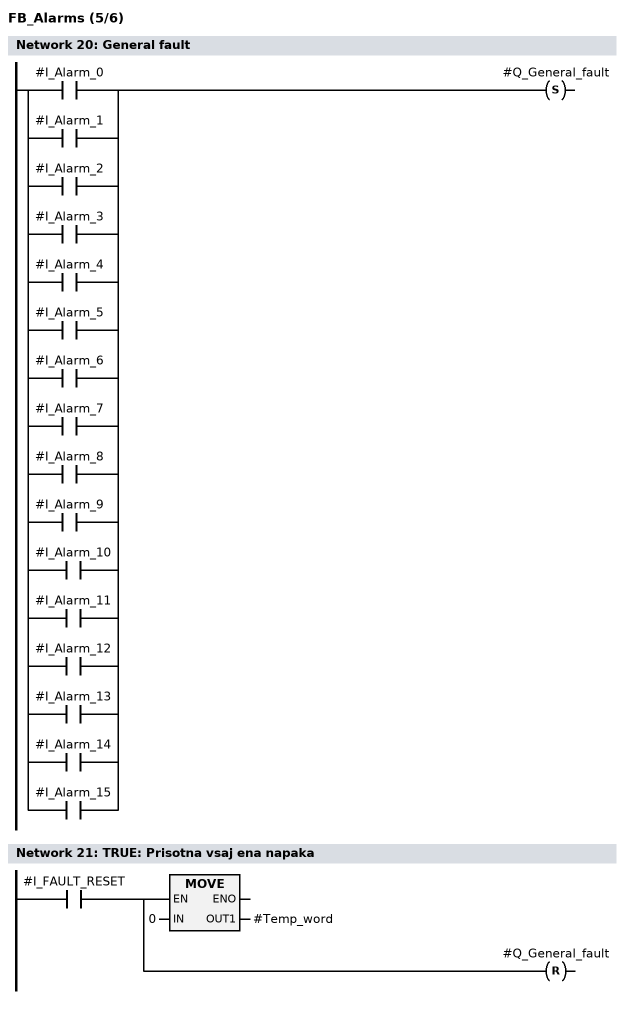
   RUNG wire#powerrail
      Contact( #I_Alarm_0 )
      wire#w1
      S_Coil( #Q_General_fault )
   END_RUNG
   RUNG wire#powerrail
      Contact( #I_Alarm_1 )
   END_RUNG wire#w1
   RUNG wire#powerrail
      Contact( #I_Alarm_2 )
   END_RUNG wire#w1
   RUNG wire#powerrail
      Contact( #I_Alarm_3 )
   END_RUNG wire#w1
   RUNG wire#powerrail
      Contact( #I_Alarm_4 )
   END_RUNG wire#w1
   RUNG wire#powerrail
      Contact( #I_Alarm_5 )
   END_RUNG wire#w1
   RUNG wire#powerrail
      Contact( #I_Alarm_6 )
   END_RUNG wire#w1
   RUNG wire#powerrail
      Contact( #I_Alarm_7 )
   END_RUNG wire#w1
   RUNG wire#powerrail
      Contact( #I_Alarm_8 )
   END_RUNG wire#w1
   RUNG wire#powerrail
      Contact( #I_Alarm_9 )
   END_RUNG wire#w1
   RUNG wire#powerrail
      Contact( #I_Alarm_10 )
   END_RUNG wire#w1
   RUNG wire#powerrail
      Contact( #I_Alarm_11 )
   END_RUNG wire#w1
   RUNG wire#powerrail
      Contact( #I_Alarm_12 )
   END_RUNG wire#w1
   RUNG wire#powerrail
      Contact( #I_Alarm_13 )
   END_RUNG wire#w1
   RUNG wire#powerrail
      Contact( #I_Alarm_14 )
   END_RUNG wire#w1
   RUNG wire#powerrail
      Contact( #I_Alarm_15 )
   END_RUNG wire#w1
   // the same network as SCL:
   IF #I_Alarm_0 OR #I_Alarm_1 OR #I_Alarm_2 OR #I_Alarm_3 OR #I_Alarm_4 OR #I_Alarm_5 OR #I_Alarm_6 OR #I_Alarm_7 OR #I_Alarm_8 OR #I_Alarm_9 OR #I_Alarm_10 OR #I_Alarm_11 OR #I_Alarm_12 OR #I_Alarm_13 OR #I_Alarm_14 OR #I_Alarm_15 THEN
       #Q_General_fault := TRUE;
   END_IF;
END_REGION

REGION Network 21: TRUE: Prisotna vsaj ena napaka
   RUNG wire#powerrail
      Contact( #I_FAULT_RESET )
      wire#w1
      { S7_GenerateENO := "TRUE" } Move(in := 0, out1 => #Temp_word)
   END_RUNG
   RUNG wire#w1
      R_Coil( #Q_General_fault )
   END_RUNG
   // the same network as SCL:
   IF #I_FAULT_RESET THEN
       #Temp_word := 0;
       #Q_General_fault := FALSE;
   END_IF;
END_REGION

REGION Network 23
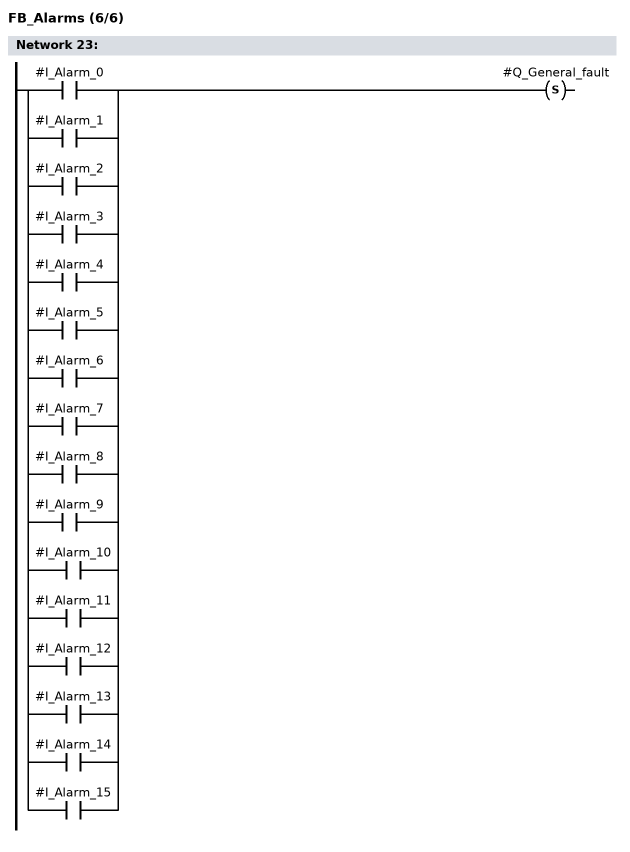
   RUNG wire#powerrail
      Contact( #I_Alarm_0 )
      wire#w1
      S_Coil( #Q_General_fault )
   END_RUNG
   RUNG wire#powerrail
      Contact( #I_Alarm_1 )
   END_RUNG wire#w1
   RUNG wire#powerrail
      Contact( #I_Alarm_2 )
   END_RUNG wire#w1
   RUNG wire#powerrail
      Contact( #I_Alarm_3 )
   END_RUNG wire#w1
   RUNG wire#powerrail
      Contact( #I_Alarm_4 )
   END_RUNG wire#w1
   RUNG wire#powerrail
      Contact( #I_Alarm_5 )
   END_RUNG wire#w1
   RUNG wire#powerrail
      Contact( #I_Alarm_6 )
   END_RUNG wire#w1
   RUNG wire#powerrail
      Contact( #I_Alarm_7 )
   END_RUNG wire#w1
   RUNG wire#powerrail
      Contact( #I_Alarm_8 )
   END_RUNG wire#w1
   RUNG wire#powerrail
      Contact( #I_Alarm_9 )
   END_RUNG wire#w1
   RUNG wire#powerrail
      Contact( #I_Alarm_10 )
   END_RUNG wire#w1
   RUNG wire#powerrail
      Contact( #I_Alarm_11 )
   END_RUNG wire#w1
   RUNG wire#powerrail
      Contact( #I_Alarm_12 )
   END_RUNG wire#w1
   RUNG wire#powerrail
      Contact( #I_Alarm_13 )
   END_RUNG wire#w1
   RUNG wire#powerrail
      Contact( #I_Alarm_14 )
   END_RUNG wire#w1
   RUNG wire#powerrail
      Contact( #I_Alarm_15 )
   END_RUNG wire#w1
   // the same network as SCL:
   IF #I_Alarm_0 OR #I_Alarm_1 OR #I_Alarm_2 OR #I_Alarm_3 OR #I_Alarm_4 OR #I_Alarm_5 OR #I_Alarm_6 OR #I_Alarm_7 OR #I_Alarm_8 OR #I_Alarm_9 OR #I_Alarm_10 OR #I_Alarm_11 OR #I_Alarm_12 OR #I_Alarm_13 OR #I_Alarm_14 OR #I_Alarm_15 THEN
       #Q_General_fault := TRUE;
   END_IF;
END_REGION
END_FUNCTION_BLOCK

FUNCTION_BLOCK "BOOL_TO_INT"   // FB125, LAD
TITLE = Alarm blok
{ S7_Optimized_Access := 'TRUE' }
AUTHOR : Andrej
VERSION : 0.1
   VAR_INPUT
      BOOL_0 : Bool;
      BOOL_1 : Bool;
      BOOL_2 : Bool;
      BOOL_3 : Bool;
      BOOL_4 : Bool;
      BOOL_5 : Bool;
      BOOL_6 : Bool;
      BOOL_7 : Bool;
      BOOL_8 : Bool;
      BOOL_9 : Bool;
      BOOL_10 : Bool;
      BOOL_11 : Bool;
      BOOL_12 : Bool;
      BOOL_13 : Bool;
      BOOL_14 : Bool;
      BOOL_15 : Bool;
   END_VAR
   VAR_OUTPUT
      "INT" : Word;
   END_VAR
   VAR RETAIN
      Temp_word : Word;
   END_VAR
BEGIN

REGION Network 1
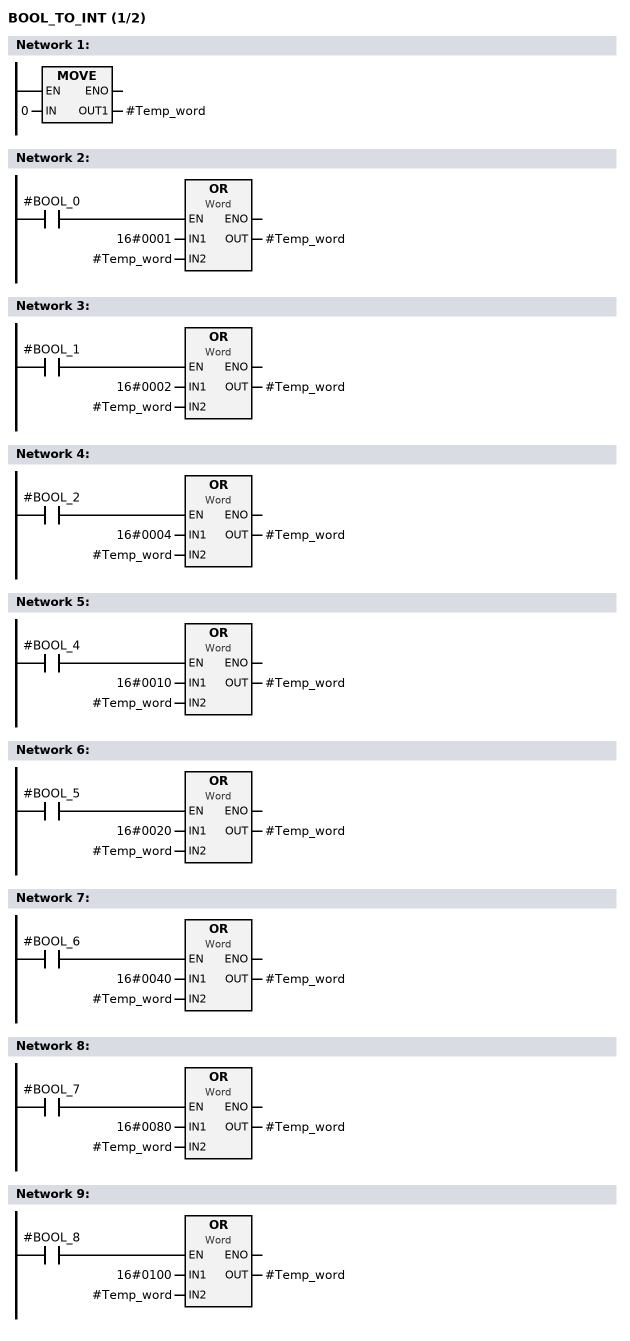
   RUNG wire#powerrail
      Move(in := 0, out1 => #Temp_word)
   END_RUNG
   // the same network as SCL:
   #Temp_word := 0;
END_REGION

REGION Network 2
   IF #BOOL_0 THEN #Temp_word := 16#0001 OR #Temp_word; END_IF;
END_REGION

REGION Network 3
   IF #BOOL_1 THEN #Temp_word := 16#0002 OR #Temp_word; END_IF;
END_REGION

REGION Network 4
   IF #BOOL_2 THEN #Temp_word := 16#0004 OR #Temp_word; END_IF;
END_REGION

REGION Network 5
   IF #BOOL_4 THEN #Temp_word := 16#0010 OR #Temp_word; END_IF;
END_REGION

REGION Network 6
   IF #BOOL_5 THEN #Temp_word := 16#0020 OR #Temp_word; END_IF;
END_REGION

REGION Network 7
   IF #BOOL_6 THEN #Temp_word := 16#0040 OR #Temp_word; END_IF;
END_REGION

REGION Network 8
   IF #BOOL_7 THEN #Temp_word := 16#0080 OR #Temp_word; END_IF;
END_REGION

REGION Network 9
   IF #BOOL_8 THEN #Temp_word := 16#0100 OR #Temp_word; END_IF;
END_REGION

REGION Network 10
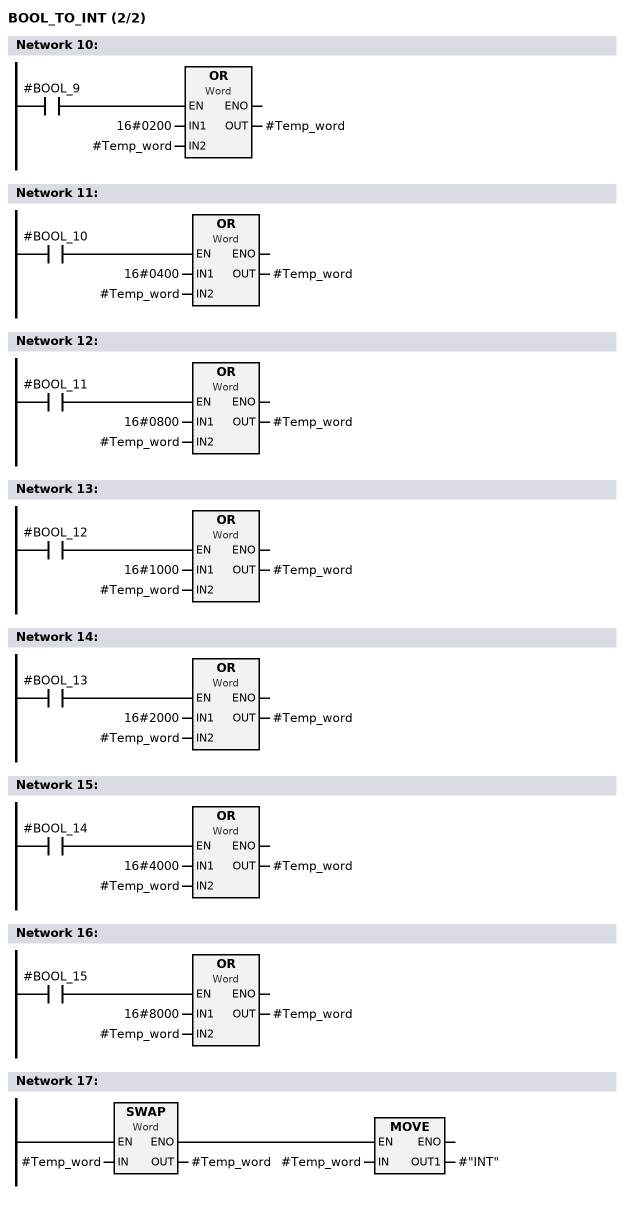
   IF #BOOL_9 THEN #Temp_word := 16#0200 OR #Temp_word; END_IF;
END_REGION

REGION Network 11
   IF #BOOL_10 THEN #Temp_word := 16#0400 OR #Temp_word; END_IF;
END_REGION

REGION Network 12
   IF #BOOL_11 THEN #Temp_word := 16#0800 OR #Temp_word; END_IF;
END_REGION

REGION Network 13
   IF #BOOL_12 THEN #Temp_word := 16#1000 OR #Temp_word; END_IF;
END_REGION

REGION Network 14
   IF #BOOL_13 THEN #Temp_word := 16#2000 OR #Temp_word; END_IF;
END_REGION

REGION Network 15
   IF #BOOL_14 THEN #Temp_word := 16#4000 OR #Temp_word; END_IF;
END_REGION

REGION Network 16
   IF #BOOL_15 THEN #Temp_word := 16#8000 OR #Temp_word; END_IF;
END_REGION

REGION Network 17
   #Temp_word := SWAP(#Temp_word);
   #"INT" := #Temp_word;
END_REGION
END_FUNCTION_BLOCK

(* ===== HMI "HMI_RT_6" =====
system functions are stored by id; their names below are inferred from use
connection "HMI_Connection_8": 
connection "HMI_Connection_1": ETHERNET, S7_1500_OMS

HMI tags "Default tag table"
   "PozKontaktNaKoncuLetve" : Bool = PLC PozKontaktNaKoncuLetve AT %I20.4, 1 s
   "FB_STARTUP_DB_korak" : UInt = PLC FB_STARTUP_DB.korak, 1 s
   "FB_IOL_IFM_SV_DB_uPretok" : UInt = PLC FB_IOL_IFM_SV_DB.uPretok, 1 s
   "FB_IOL_IFM_SV_DB_fTemperatura" : Real = PLC FB_IOL_IFM_SV_DB.fTemperatura, 1 s
   "FB_FESTO_VPPM_DB_TrenutniPritisk" : Real = PLC FB_FESTO_VPPM_DB.TrenutniPritisk, 1 s
   "FB_FESTO_SDE1_DB_oPritisk" : Real = PLC FB_FESTO_SDE1_DB.oPritisk, 1 s
   "FB_Lin_FESTO_PNEVMATIKA_PRITISK_Q_izhod" : Real = PLC FB_Lin_FESTO_PNEVMATIKA_PRITISK.Q_izhod, 1 s
   "FB_FESTO_VPPM_DB_setstatZeljeniPritisk" : Real = PLC FB_FESTO_VPPM_DB.setstatZeljeniPritisk, 1 s
   "Keyence_OdmičniCilinderKonusa" : DInt = PLC Keyence_OdmičniCilinderKonusa AT %ID137, 1 s
   "Keyence_OdmičniCilinderVarjenja" : DInt = PLC Keyence_OdmičniCilinderVarjenja AT %ID144, 1 s
   "DB_HMI_ROČNI NAČIN_izbraniCilinder" : Int = PLC DB_HMI."ROČNI NAČIN".izbraniCilinder, 1 s
   "ZaporaIzdelka" : Bool = PLC ZaporaIzdelka AT %I20.0, 1 s
   "SprositevZaporeIzdelka" : Bool = PLC SprositevZaporeIzdelka AT %I20.1, 1 s
   "1Y1_OdklepZapore" : Bool = PLC 1Y1_OdklepZapore AT %Q44.0, 1 s
   "Y2/1_NalaganjeNazanj" : Bool = PLC "Y2/1_NalaganjeNazanj" AT %Q44.3, 1 s
   "Y2/1_NalaganjeNaprej" : Bool = PLC "Y2/1_NalaganjeNaprej" AT %Q44.2, 1 s
   "DB_HMI_SDAT1_PozPobiranje" : Real = PLC DB_HMI.SDAT1.PozPobiranje, 1 s
   "DB_HMI_SDAT1_PozNalaganje" : Real = PLC DB_HMI.SDAT1.PozNalaganje, 1 s
   "SDAT1_oPoz1Dosezena" : Bool = PLC SDAT1.oPoz1Dosezena, 1 s
   "SDAT2_oPoz2Dosezena" : Bool = PLC SDAT2.oPoz2Dosezena, 1 s
   "SDAT1_oPoz2Dosezena" : Bool = PLC SDAT1.oPoz2Dosezena, 1 s
   "Y3/1_PrijemaloKontaktaOdpri" : Bool = PLC "Y3/1_PrijemaloKontaktaOdpri" AT %Q44.4, 1 s
   "PrijemaloKontaktaOdprto" : Bool = PLC PrijemaloKontaktaOdprto AT %I20.3, 1 s
   "PrijemaloKontaktaZaprto" : Bool = PLC PrijemaloKontaktaZaprto AT %I20.2, 1 s
   "DB_HMI_SDAT2_PozNalaganje" : Real = PLC DB_HMI.SDAT2.PozPobiranjePloscice, 1 s
   "DB_HMI_SDAT2_PozPobiranje" : Real = PLC DB_HMI.SDAT2.PozNalaganjePloscice, 1 s
   "SDAT1_out" : Real = PLC SDAT1.out, 1 s
   "SDAT2_out" : Real = PLC SDAT2.out, 1 s
   "FB_KEYENCE_GT2_ODMIKVARJENJA_oPoz1Dosezena" : Bool = PLC FB_KEYENCE_GT2_ODMIKVARJENJA.oPoz1Dosezena, 1 s
   "FB_KEYENCE_GT2_ODMIKVARJENJA_oPoz3Dosezena" : Bool = PLC FB_KEYENCE_GT2_ODMIKVARJENJA.oPoz3Dosezena, 1 s
   "Y1/3_odmičniCilinderVarjenje_GOR" : Bool = PLC "Y1/4_odmičniCilinderVarjenje_GOR" AT %Q46.4, 1 s
   "Y1/3_odmičniCilinderVarjenjeDOL" : Bool = PLC "Y1/4_odmičniCilinderVarjenjeDOL" AT %Q46.5, 1 s
   "PozKontaktNazaj" : Bool = PLC PozKontaktNazaj AT %I20.7, 1 s
   "PozKontaktNaprej" : Bool = PLC PozKontaktNaprej AT %I20.6, 1 s
   "Y2/3_PozicioniranjeKontaktovNazaj" : Bool = PLC "Y2/3_PozicioniranjeKontaktovNazaj" AT %Q45.2, 1 s
   "Y2/3_PozicioniranjeKontaktovNaprej" : Bool = PLC "Y2/3_PozicioniranjeKontaktovNaprej" AT %Q45.3, 1 s
   "Y1/3_OdmičniCilinderKonusa" : Bool = PLC "Y1/3_OdmičniCilinderKonusa" AT %Q45.0, 1 s
   "DB_KEYENCE_Kroznik_ZeljenaPozicija_POZ1" : UInt = PLC DB_KEYENCE.Kroznik.ZeljenaPozicija.POZ1_KonusNazaj, 1 s
   "DB_KEYENCE_Kroznik_ZeljenaPozicija_POZ2" : UInt = PLC DB_KEYENCE.Kroznik.ZeljenaPozicija.POZ2_KonusNaprej, 1 s
   "FB_KEYENCE_GT2_odmikKonusaKroznika_oPoz1Dosezena" : Bool = PLC FB_KEYENCE_GT2_odmikKonusaKroznika.oPoz1Dosezena, 1 s
   "FB_KEYENCE_GT2_odmikKonusaKroznika_oPoz2Dosezena" : Bool = PLC FB_KEYENCE_GT2_odmikKonusaKroznika.oPoz2Dosezena, 1 s
   "DrzanjeKontakta" : Bool = PLC DrzanjeKontakta AT %I21.1, 1 s
   "Y3/3_OdpiranjeDržalaKomada" : Bool = PLC "Y3/3_OdpiranjeDržalaKomada" AT %Q45.4, 1 s
   "Y4/3_OdpiranjeIzmetaKontakta" : Bool = PLC "Y4/3_OdpiranjeIzmetaKontakta" AT %Q45.6, 1 s
   "DrzanjeIzmetKontakta" : Bool = PLC DrzanjeIzmetKontakta AT %I21.0, 1 s
   "IzmetKontaktaNazaj" : Bool = PLC IzmetKontaktaNazaj AT %I21.2, 1 s
   "Y5/3_IzmetKomadov" : Bool = PLC "Y5/3_IzmetKomadov" AT %Q46.0, 1 s
   "DrscaSLabiKosi" : Bool = PLC DrscaSLabiKosi AT %I21.5, 1 s
   "DrcaDobriKosi" : Bool = PLC DrcaDobriKosi AT %I21.4, 1 s
   "Y6/3_LoputaSlabi" : Bool = PLC "Y6/3_LoputaSlabi" AT %Q46.3, 1 s
   "Y6/3_LoputaDobri" : Bool = PLC "Y6/3_LoputaDobri" AT %Q46.2, 1 s
   "DB_KEYENCE_Elektroda_ZeljenaPozicija_POZ1" : UInt = PLC DB_KEYENCE.Elektroda.ZeljenaPozicija.POZ1_elektrodaGor, 1 s
   "DB_KEYENCE_Elektroda_ZeljenaPozicija_POZ2" : UInt = PLC DB_KEYENCE.Elektroda.ZeljenaPozicija.POZ2_elektrodaVmes, 1 s
   "DB_KEYENCE_Elektroda_ZeljenaPozicija_POZ3_elektrodaStisnjena" : UInt = PLC DB_KEYENCE.Elektroda.ZeljenaPozicija.POZ3_elektrodaStisnjena, 1 s
   "DB_KEYENCE_Elektroda_ZeljenaPozicija_POZ4_elektrodaZavarjeno" : UInt = PLC DB_KEYENCE.Elektroda.ZeljenaPozicija.POZ4_elektrodaZavarjeno, 1 s
   "FB_KEYENCE_GT2_ODMIKVARJENJA_oPoz2Dosezena" : Bool = PLC FB_KEYENCE_GT2_ODMIKVARJENJA.oPoz2Dosezena, 1 s
   "FB_KEYENCE_GT2_ODMIKVARJENJA_oPoz4Dosezena" : Bool = PLC FB_KEYENCE_GT2_ODMIKVARJENJA.oPoz4Dosezena, 1 s
   "Y2_1_dovajanjeKntaktovNaprej" : Bool = PLC Y2_1_dovajanjePlosciceNaprej AT %Q44.7, 1 s
   "Y2/1_dovajanjeKontaktovNazaj" : Bool = PLC "Y2/1_dovajanjePlosciceNazaj" AT %Q44.6, 1 s
   "RežimDelovanja" : Byte = PLC RežimDelovanja AT %MB3, 1 s
   "FB_Alarms_DB_Q_Alarm_word" : Word = PLC FB_Alarms_DB.Q_Alarm_word, 1 s
   "DB_PODATKI_GeaphName" : String[254] = PLC DB_PODATKI.GeaphName, 1 s
   "GRAPH_HMI_HMINAME{0}" : String[254] = PLC GRAPH_HMI.HMINAME[0] AT %DB38.DBX0.0, 1 s
   "SDAT2_oPoz1Dosezena" : Bool = PLC SDAT2.oPoz1Dosezena, 1 s
   "FB_STARTUP_DB_DeviceState_mySTATE{7}" : Bool = PLC FB_STARTUP_DB.DeviceState.mySTATE[7], 1 s
   "FB_STARTUP_DB_DeviceState_mySTATE{8}" : Bool = PLC FB_STARTUP_DB.DeviceState.mySTATE[8], 1 s
   "FB_AKD_Kroznik_iAKD_PODATKI_TO_SIEMENS_HomePosSet" : Bool = PLC FB_AKD_Kroznik.iAKD.PODATKI_TO_SIEMENS.HomePosSet, 1 s
   "FB_AKD_Kroznik_iAKD_PODATKI_TO_SIEMENS_FaultPresent" : Bool = PLC FB_AKD_Kroznik.iAKD.PODATKI_TO_SIEMENS.FaultPresent, 1 s
   "FB_AKD_VrtenjeELektrode_iAKD_PODATKI_TO_SIEMENS_ErrInRange" : Bool = PLC FB_AKD_VrtenjeELektrode.iAKD.PODATKI_TO_SIEMENS.ErrInRange, 1 s
   "FB_AKD_VrtenjeELektrode_iAKD_PODATKI_TO_SIEMENS_HomePosSet" : Bool = PLC FB_AKD_VrtenjeELektrode.iAKD.PODATKI_TO_SIEMENS.HomePosSet, 1 s
   "FB_STARTUP_DB_DeviceState_mySTATE{5}" : Bool = PLC FB_STARTUP_DB.DeviceState.mySTATE[5], 1 s
   "FB_AKD_REZANJEPODAJANJE_iAKD_PODATKI_TO_SIEMENS_FaultPresent" : Bool = PLC FB_AKD_REZANJEPODAJANJE.iAKD.PODATKI_TO_SIEMENS.FaultPresent, 1 s
   "FB_AKD_REZANJEPODAJANJE_iAKD_PODATKI_TO_SIEMENS_HomePosSet" : Bool = PLC FB_AKD_REZANJEPODAJANJE.iAKD.PODATKI_TO_SIEMENS.HomePosSet, 1 s
   "FB_AKD_DB_elektroda_iAKD_PODATKI_TO_SIEMENS_FaultPresent" : Bool = PLC FB_AKD_DB_elektroda.iAKD.PODATKI_TO_SIEMENS.FaultPresent, 1 s
   "FB_AKD_DB_RezanjePodajanje_iAKD_PODATKI_TO_SIEMENS_FaultPresent" : Bool = PLC FB_AKD_DB_RezanjePodajanje.iAKD.PODATKI_TO_SIEMENS.FaultPresent, 1 s
   "TimerReady" : Bool = PLC TimerReady AT %I66.3, 1 s
   "WeldFault" : Bool = PLC WeldFault AT %I66.4, 1 s
   "EndOfSequency_WC" : Bool = PLC EndOfSequency_WC AT %I66.2, 1 s
   "FB_IOL_IFM_SV_DB_oPretokOK" : Bool = PLC FB_IOL_IFM_SV_DB.oPretokOK, 1 s
   "FB_IOL_IFM_SV_DB_oTempOK" : Bool = PLC FB_IOL_IFM_SV_DB.oTempOK, 1 s
   "ExternalWeldOn" : Bool = PLC ExternalWeldOn AT %Q53.0, 1 s
   "DB_PODATKI_KROZNA_MIZA_IzdelekPrisoten" : Byte = PLC DB_PODATKI.KROZNA_MIZA.IzdelekPrisoten, 500 ms
   "DB_PODATKI_KROZNA_MIZA_IzdelekPrisotenArray{7}" : Bool = PLC DB_PODATKI.KROZNA_MIZA.IzdelekPrisotenArray[7], 100 ms
   "DB_PODATKI_KROZNA_MIZA_StatusIzdelka{7}" : Byte = PLC DB_PODATKI.KROZNA_MIZA.StatusIzdelkaVarjenje[7], 100 ms
   "DB_PODATKI_KROZNA_MIZA_StatusIzdelka{6}" : Byte = PLC DB_PODATKI.KROZNA_MIZA.StatusIzdelkaVarjenje[6], 100 ms
   "DB_PODATKI_KROZNA_MIZA_StatusIzdelka{5}" : Byte = PLC DB_PODATKI.KROZNA_MIZA.StatusIzdelkaVarjenje[5], 100 ms
   "DB_PODATKI_KROZNA_MIZA_StatusIzdelka{4}" : Byte = PLC DB_PODATKI.KROZNA_MIZA.StatusIzdelkaVarjenje[4], 500 ms
   "DB_PODATKI_KROZNA_MIZA_StatusIzdelka{3}" : Byte = PLC DB_PODATKI.KROZNA_MIZA.StatusIzdelkaVarjenje[3], 500 ms
   "DB_PODATKI_KROZNA_MIZA_StatusIzdelka{2}" : Byte = PLC DB_PODATKI.KROZNA_MIZA.StatusIzdelkaVarjenje[2], 500 ms
   "FB_Alarms_DB_1_Q_Alarm_word" : Word = PLC FB_Alarms_DB_1.Q_Alarm_word, 1 s
   "DB_PODATKI_KROZNA_MIZA_IzdelekPrisotenArray{5}" : Bool = PLC DB_PODATKI.KROZNA_MIZA.IzdelekPrisotenArray[5], 100 ms
   "DB_PODATKI_KROZNA_MIZA_IzdelekPrisotenArray{4}" : Bool = PLC DB_PODATKI.KROZNA_MIZA.IzdelekPrisotenArray[4], 500 ms
   "DB_PODATKI_KROZNA_MIZA_IzdelekPrisotenArray{3}" : Bool = PLC DB_PODATKI.KROZNA_MIZA.IzdelekPrisotenArray[3], 500 ms
   "DB_PODATKI_KROZNA_MIZA_IzdelekPrisotenArray{2}" : Bool = PLC DB_PODATKI.KROZNA_MIZA.IzdelekPrisotenArray[2], 500 ms
   "DB_PODATKI_KROZNA_MIZA_IzdelekPrisotenArray{1}" : Bool = PLC DB_PODATKI.KROZNA_MIZA.IzdelekPrisotenArray[1], 100 ms
   "DB_PODATKI_KROZNA_MIZA_StatusIzdelkaVarjenje{1}" : Byte = PLC DB_PODATKI.KROZNA_MIZA.StatusIzdelkaVarjenje[1], 100 ms
   "FB_AKD_Kroznik_iAKD_PODATKI_TO_SIEMENS_WarningPreent" : Bool = PLC FB_AKD_Kroznik.iAKD.PODATKI_TO_SIEMENS.WarningPreent, 1 s
   "FB_AKD_VrtenjeELektrode_iAKD_PODATKI_TO_SIEMENS_WarningPreent" : Bool = PLC FB_AKD_VrtenjeELektrode.iAKD.PODATKI_TO_SIEMENS.WarningPreent, 1 s
   "FB_AKD_REZANJEPODAJANJE_iAKD_PODATKI_TO_SIEMENS_WarningPreent" : Bool = PLC FB_AKD_REZANJEPODAJANJE.iAKD.PODATKI_TO_SIEMENS.WarningPreent, 1 s
   "DB_UDP_COMM_PLC_TO_PC_TUSEND_DB_TUSEND_REQ" : Bool = PLC DB_UDP_COMM.PLC_TO_PC.TUSEND_DB.TUSEND_REQ AT %DB17.DBX1044.0, 1 s
   "PrisotnostTraka" : Bool = PLC PrisotnostTraka AT %I8.6, 1 s
   "FB_AKD_DB_elektroda_o_BerrStatus" : Byte = PLC FB_AKD_DB_elektroda.o_BerrStatus, 1 s
   "FB_AKD_Kroznik_o_BerrStatus" : Byte = PLC FB_AKD_Kroznik.o_BerrStatus, 1 s
   "FB_AKD_DB_RezanjePodajanje_o_BerrStatus" : Byte = PLC FB_AKD_DB_RezanjePodajanje.o_BerrStatus, 1 s
   "DB_PODATKI_KROZNA_MIZA_IzdelekPrisotenArray{6}" : Bool = PLC DB_PODATKI.KROZNA_MIZA.IzdelekPrisotenArray[6], 100 ms
   "FB_AKD_Kroznik_bPogojiZaVKLOP" : Bool = PLC FB_AKD_Kroznik.bPogojiZaVKLOP, 1 s
   "FB_AKD_DB_elektroda_bPogojiZaVKLOP" : Bool = PLC FB_AKD_DB_elektroda.bPogojiZaVKLOP, 1 s
   "STEVEC_KOSOV" : Counter = PLC STEVEC_KOSOV AT %C0, 1 s
   "DB_KEYENCE_Elektroda_TOLERANCA{1}" : Int = PLC DB_KEYENCE.Elektroda.TOLERANCA[1], 1 s
   "DB_KEYENCE_Elektroda_TOLERANCA{2}" : Int = PLC DB_KEYENCE.Elektroda.TOLERANCA[2], 1 s
   "DB_KEYENCE_Elektroda_TOLERANCA{3}" : Int = PLC DB_KEYENCE.Elektroda.TOLERANCA[3], 1 s
   "DB_KEYENCE_Elektroda_TOLERANCA{4}" : Int = PLC DB_KEYENCE.Elektroda.TOLERANCA[4], 1 s
   "DB_KEYENCE_TOLERANCA{1}" : Int = PLC DB_KEYENCE.TOLERANCA[1], 1 s
   "DB_KEYENCE_TOLERANCA{2}" : Int = PLC DB_KEYENCE.TOLERANCA[2], 1 s
   "GraphTab" : WString[10], internal
   "StatusCode" : Byte = PLC StatusCode AT %IB82, 1 s
   "DB_HMI_Varjenje_ResetWithWC" : Bool = PLC DB_HMI.Varjenje.ResetWithWC, 1 s
   "FB_AKD_VrtenjeKroznika_o_BerrStatus" : Byte = PLC FB_AKD_VrtenjeKroznika.o_BerrStatus, 1 s
   "StatusPrisotnostiTraku" : Byte = PLC StatusPrisotnostiTraku AT %MB5, 1 s
   "NapakaOdvijanjaTrau" : Bool = PLC NapakaOdvijanjaTrau AT %M4.2, 1 s
   "NapakaCiscenjaElektrode" : Bool = PLC NapakaCiscenjaElektrode AT %M4.3, 1 s
   "DB_STEVCI_STEVCI_SKUPAJ" : UInt = PLC DB_STEVCI."STEVCI VARJENJE".SKUPAJ, 1 s
   "db_AKD_REZANJEPODAJANJE_PODATKI_PloscicaOdrezana" : Bool = PLC db_AKD.REZANJEPODAJANJE.PODATKI.PloscicaOdrezana, 1 s
   "DB_STEVCI_STEVCI_SKUPAJOK" : UInt = PLC DB_STEVCI."STEVCI VARJENJE".SKUPAJOK, 1 s
   "DB_STEVCI_STEVCI_ZavarjenoOK" : UInt = PLC DB_STEVCI."STEVCI VARJENJE".ZavarjenoOK, 1 s
   "DB_STEVCI_STEVCI_ZavarjenoNOK" : UInt = PLC DB_STEVCI."STEVCI VARJENJE".ZavarjenoNOK, 1 s
   "DB_STEVCI_STEVCI KAMERA_SKUPAJ" : UInt = PLC DB_STEVCI."STEVCI KAMERA".SKUPAJ, 1 s
   "DB_STEVCI_STEVCI KAMERA_KameraOK" : UInt = PLC DB_STEVCI."STEVCI KAMERA".KameraOK, 1 s
   "DB_STEVCI_STEVCI KAMERA_KameraNOK" : UInt = PLC DB_STEVCI."STEVCI KAMERA".KameraNOK, 1 s
   "DB_STEVCI_STEVEC_SKATEL_SKATLA1" : UInt = PLC DB_STEVCI.STEVEC_SKATEL.SKATLA1, 1 s
   "DB_STEVCI_STEVEC_SKATEL_SKATLA2" : UInt = PLC DB_STEVCI.STEVEC_SKATEL.SKATLA2, 1 s
   "Clock_1Hz" : Bool = PLC Clock_1Hz AT %M0.5, 500 ms
   "DB_HMI_TekočiTrak_btnResetSkatle1" : Bool = PLC DB_HMI.TekočiTrak.btnResetSkatle1, 1 s
   "DB_HMI_TekočiTrak_btnResetSKatle2" : Bool = PLC DB_HMI.TekočiTrak.btnResetSKatle2, 1 s
   "DB_STEVCI_STEVCI_ZELENAPOLNA_SKATLA_SKATLA1" : UInt = PLC DB_STEVCI.STEVCI_ZELENAPOLNA_SKATLA.SKATLA1, 1 s
   "DB_STEVCI_STEVCI_ZELENAPOLNA_SKATLA_SKATLA2" : UInt = PLC DB_STEVCI.STEVCI_ZELENAPOLNA_SKATLA.SKATLA2, 1 s
   "FB_TekociTrak_DB_stat_skatla1Polna" : Bool = PLC FB_TekociTrak_DB.stat_skatla1Polna, 1 s
   "FB_TekociTrak_DB_stat_skatla2Polna" : Bool = PLC FB_TekociTrak_DB.stat_skatla2Polna, 1 s
   "db_AKD_KROZNIK_PODATKI_StartHomming" : Bool = PLC db_AKD.KROZNIK.PODATKI.StartHomming, 1 s
   "DB_HMI_Kroznik_bStartHomming" : Bool = PLC DB_HMI.Kroznik.bStartHomming, 1 s
   "FB_AKD_VrtenjeKroznika_iAKD_PODATKI_TO_SIEMENS_HomePosSet" : Bool = PLC FB_AKD_VrtenjeKroznika.iAKD.PODATKI_TO_SIEMENS.HomePosSet, 1 s
   "FB_AKD_VrtenjeKroznika_OmogociHome" : Bool = PLC FB_AKD_VrtenjeKroznika.OmogociHome, 1 s
   "SenzorOdvijanjaCiscenjeElektrode" : Bool = PLC SenzorOdvijanjaCiscenjeElektrode AT %I21.6, 1 s
   "FB_CYCLETIME_cycleTime" : LTime = PLC FB_CYCLETIME.cycleTime, 1 s
   "FB_CYCLETIME_CycleTimeTIe" : Time = PLC FB_CYCLETIME.CycleTimeTIe, 1 s
   "FB_CYCLETIME_TimeReal" : Real = PLC FB_CYCLETIME.TimeReal, 1 s
   "FB_CYCLETIME_IzdelkiNaUro" : Int = PLC FB_CYCLETIME.IzdelkiNaUro, 1 s
   "FB_CYCLETIME_mm" : Int = PLC FB_CYCLETIME.mm, 1 min
   "DB_HMI_HMI_izpisNapak_w_trenutnaNapak" : WString[254] = PLC DB_HMI.HMI_izpisNapak.w_trenutnaNapak, 1 s
   "WSTR_HMI_NAPAKA" : WString[254] = PLC DB_HMI.HMI_izpisNapak.w_trenutnaNapak, 1 s
   "HMI_Tag_1" : WString[10], internal
   "DB_HMI_ČiščenjeElektrode_ZeljenoStevilo" : UInt = PLC DB_HMI.ČiščenjeElektrode.ZeljenoStevilo, 1 s
   "FB_CYCLETIME_staticmm" : Int = PLC FB_CYCLETIME.staticmm, 1 s
   "FB_CYCLETIME_intfloor" : Int = PLC FB_CYCLETIME.intfloor, 1 s
   "Clock_2.5Hz" : Bool = PLC "Clock_2.5Hz" AT %M0.2, 1 s
   "Clock_5Hz" : Bool = PLC Clock_5Hz AT %M0.1, 100 ms
      on ChangeValue: "VBFunction_1"()
   "FB_LocalTime_DB_DateAndTIME" : LDT = PLC FB_LocalTime_DB.DateAndTIME, 1 s
   "FB_LocalTime_DB_WR_LOC_LOCALTIME" : LDT = PLC FB_LocalTime_DB.WR_LOC.LOCALTIME, 1 s
   "FB_KAMERA_TRIG_DB_stat_CamLastValue" : Bool = PLC FB_KAMERA_TRIG_DB.stat_CamLastValue, 1 s
   "FB_KAMERA_TRIG_DB_io_StatusArrayCamere" : Byte = PLC FB_KAMERA_TRIG_DB.io_StatusArrayCamere, 1 s

HMI tags "Template"
   "MainNavigationState" : Int, internal
   "SubNavigationState" : Int, internal
   "CurrentUserName" : WString[18], internal
   "DiagState" : Int, internal
   "PopUpBackground" : Bool, internal
   "UserName" : WString[20], internal
   "Password" : WString[20], internal
   "UserIsLoggedIn" : Bool, internal
   "CodeView" : Bool, internal
   "Brightness" : Int, internal
   "CurrentLanguage" : Bool, internal
   "CurrentRecipeName" : WString[30], internal
   "CurrentMachineState" : Int, internal
   "OptionPanelNavigationState" : Int, internal
   "ButtonDown" : Bool, internal
   "ThirdLevelNavigationState" : Int, internal
   "StartScreenName" : WString[60], internal
   "InScreenTabState" : Int, internal
   "DummyTagBool" : Bool, internal
   "DummyTagInt1" : Int, internal
   "DummyTagInt2" : Int, internal
   "DummyTagInt3" : Int, internal
   "DummyDeltaReal" : LReal, internal
   "DummTagReal1" : LReal, internal
   "DummyDeltaInt" : Int, internal

discrete alarms
   2: 'Pozicija pred varjenjem neustrezna / Preveri ali je ploščica ustrezno vstavljena', class Errors, trigger "FB_Alarms_DB_1_Q_Alarm_word" bit 0
   1: 'Premalo zraka v sistemu / Preveri dovod zraka. Preveri ali je ventil odprt.', class Errors, trigger "FB_Alarms_DB_1_Q_Alarm_word" bit 1
   3: 'Pozicija pobiranja izdelka P1 / Preveri nastavitve pozicije za pobiranje izdelka iz lin. traka', class Errors, trigger "FB_Alarms_DB_1_Q_Alarm_word" bit 2

text list "Machine State": 0 'Undefined / Kein Job'; 1 'Production / Produktion'; 2 'Startup / Anlauf'; 3 'Paused / Pausiert'; 4 'Stopped / Gestoppt'; 5 'Shutdown / Beenden'; 6 'Undefined / UNBEKANNT'; 10 'ROČNO'; 11 'AVTO'

text list "timeRange": 1 'Hours / Stunden'; 2 'Days / Tage'; 3 'Weeks / Wochen'; 4 'Months / Monate'; 5 'Years / Jahre'

text list "MachineState_Farfield": 0..1 '???'; 1 'OK'; 2 'ERROR / FEHLER'; 3 'PAUSED / HALT'

text list "Foil Types": 0..1 '120 - 1mm - Transparent'; 1 '120 - 3mm - Transparent'; 2 '240 - 1mm - Transparent'; 3 '240 - 3mm - Transparent'

text list "FunctionState": 0 'Disabled / Deaktiviert'; 1 'Enabled / Aktiviert'

text list "GroundPos": 0 'No / Nein'; 1 'Yes / Ja'

text list "State": 0 'Off / Aus'; 1 'On / An'

text list "TestiranjeStroja": 0 'Zagon PLC krmilnika...'; 5 'profinet komunikacije neuspešna'; 10 'ERROR | profinet komunikacija SIEMENS <---> MVK1 - IOL master'; 15 'ERROR | profinet komunikacija SIEMENS <---> MVK2 - IOL master'; 1 'HMI komunikacije neuspešna'; 20 'ERROR | profinet komunikacija SIEMENS <---> MVK3 - IOL master'; 25 'ERROR | profinet komunikacija z Kollmorgen AKD - cilinder'; 30 'ERROR | Profinet komunikacije z Kollmorgen AKD - vrtljiva miza'; 35 'ERROR | Profinet komunikacija z Kollmorgen AKD - elektroda'; 40 'ERROR | Profinet komunikacija z varilnikom - Bosh neuspešna'; 45 'ERROR | Profinet komunikacije z Keyence PN neuspešna'

text list "BOSH": 0 'OK'; 80 'IZKLOP_V_SILI'; 81 'WELD_WITHOUD_COMMAND'; 85 'MEMMORY_DELETED'; 87 'NO_WELDING_PROGRAM'; 91 'MAIN_SWITCH_TRIPPED'; 99 'WELD_PROCESS_ERROR'; 160 'MAX_HEAT_SINK_TEMP'

text list "StatusSkatel": 0 'OK'; 1 'Potrebna potrditev'

graphic list "DiagState": 0 'DiagOkay'; 1 'DiagWarning_1'; 2 'DiagDefault'

graphic list "DiagState_1": 0 'DiagOkay_1'; 1 'DiagWarning'; 2 'DiagDefault'

graphic list "DiagState_2": 0 'DiagOkay_1'; 1 'DiagWarning'; 2 'DiagDefault'

graphic list "DiagState_3": 0 'DiagOkay_White'; 1 'DiagWarning_White'; 2 'Circle'

graphic list "State": 0..1 'OK'; 3 'Error'

graphic list "Machine": 1 'Grafik_Verpackung_Step1_Blink-off'; 2 'Grafik_Verpackung_Step2'; 3 'Grafik_Verpackung_Blink-on'; 6..7 'Grafik_Verpackung_Step1_Blink-off'

screen "10_Start" 1280x800, template "04_PLC_StartUP"
   on GenerateScreen: "GetStartScreenName"(); "CheckCurrentUserName"()
   GraphicView "Graphic view_1" at 292,228 size 546x153; Picture "HMI_Template_Suite_Logo_Panel"
   TextField "Text field_1" at 292,492 size 343x28; Text 'Testiranje parametrov stroja...'
   SymbolicIOField "Symbolic I/O field_1" at 284,531 size 711x34; TextOff '0'; TextOn '1'; TextList "TestiranjeStroja"
      ProcessValue <- "FB_STARTUP_DB_korak"
   GraphicView "Graphic view_2" at 0,0 size 1280x800; Picture "PopUpBackground"
      Visibility <- "PopUpBackground"

screen "20_Messages" 1280x800, template "01_One_Nav_Level"
   AlarmView "Alarm view_1" at 0,104 size 1280x695
   GraphicView "Graphic view_2" at 0,0 size 1280x800; Picture "PopUpBackground"
      Visibility <- "PopUpBackground"

screen "30_Diagnostics" 1280x800, template "01_One_Nav_Level"
   SysDiagControl "System diagnostics view_1" at 0,104 size 1280x695
   GraphicView "Graphic view_2" at 0,0 size 1280x800; Picture "PopUpBackground"
      Visibility <- "PopUpBackground"

screen "40_Settings" 1280x800, template "02_Settings"
   Slider "Template_Slider_1" at 320,197 size 300x30; Caption 'SIMATIC'
      on Change: function_e4c2bb66("Brightness")
      ProcessValue <- "Brightness"
   TextField "Template_Text field_1" at 180,200 size 92x24; Text 'Brightness / Helligkeit'
   GraphicView "Graphic view_2" at 0,0 size 1280x800; Picture "PopUpBackground"
      Visibility <- "PopUpBackground"

Template "01_One_Nav_Level" 1280x800
   Gauge "gaugeDiagStateUpdate" at 566,2 size 50x50; CaptionText 'SIMATIC'
      on Change: "CheckDiagState"()
      ProcessValue <- "@DiagnosticsIndicatorTag"
   TextField "txtTitleBar" at 16,8 size 613x32; Text 'LINIJA ETI C 25 / Applikation'
   GraphicView "gfxNavigationIcon" at 1241,15 size 23x19; Picture "Hamburger_Icon"
   Button "btnNavigation" at 1224,0 size 56x48; TextOff 'Text'
      on Click: function_cf6f4242("GraphX_Slidein_Right", 1)
   Button "btnStartscreen" at 0,2 size 387x45; TextOff 'Text'
      on Click: "ActivateStartScreen"()
   TextField "txtStateHeadline" at 79,55 size 175x23; Text 'Režim vodenja stroja / Status'
   TextField "txtOperatorHeadline" at 527,55 size 129x23; Text 'Uporabnik / Bediener'
   SymbolicIOField "ioState" at 100,72 size 119x30; TextOn '1'; TextOff '0'; TextList "Machine State"
      ProcessValue <- "RežimDelovanja"
   IOField "ioOperator" at 527,72 size 126x30; FormatPattern ??????????????????
      ProcessValue <- "CurrentUserName"
   Rectangle "rectState" at 0,46 size 56x56
      Appearance <- "CurrentMachineState"
   Rectangle "rectSystemDiagnosticsIndicator" at 1224,48 size 56x56
      Appearance <- "DiagState"
   GraphicIOField "gioDiagState" at 1236,60 size 32x32; PictureList "DiagState_3"
      ProcessValue <- "DiagState"
   Button "btnDiagState" at 1224,48 size 56x56; TextOff 'Text'
      on Click: ActivateScreen("30_Diagnostics", 0)
   Button "btnOperator" at 669,56 size 40x40; TextOff '...'; PictureOff "More_Icon"
      on Click: "ShowLoginPopUp"()
   DateTimeField "Template_Date/time field_1" at 1083,64 size 133x30
      ProcessValue <- "FB_LocalTime_DB_DateAndTIME"

Template "02_Two_Nav_Levels" 1280x800
   GraphicView "gfxPrevScreenIcon" at 1240,763 size 24x24; Picture "PrevScreen_Icon"
   Button "btnSubNav1" at 0,752 size 144x48; TextOff 'Overview / Übersicht'
      on Click: SetTag("SubNavigationState", 1)
   Button "btnSubNav2" at 144,752 size 144x48; TextOff 'Module 1 / Modul 1'
      on Click: SetTag("SubNavigationState", 2)
   Button "btnSubNav3" at 288,752 size 144x48; TextOff 'Module 2 / Modul 2'
      on Click: SetTag("SubNavigationState", 3)
   Button "btnSubNav4" at 432,752 size 144x48; TextOff 'Module 3 / Modul 3'
      on Click: SetTag("SubNavigationState", 4)
   Button "btnSubNav5" at 576,752 size 144x48; TextOff 'Module 4 / Modul 4'
      on Click: SetTag("SubNavigationState", 5)
   Button "btnSubNav6" at 720,752 size 144x48; TextOff 'Module 5 / Modul 5'
      on Click: SetTag("SubNavigationState", 6)
   Button "btnSubNav7" at 864,752 size 144x48; TextOff 'Module 6 / Modul 5'
      on Click: SetTag("SubNavigationState", 7)
   Button "btnPreviousScreen" at 1224,751 size 56x48; TextOff 'Text'
      on Click: function_efd93a16()
   Gauge "gaugeDiagStateUpdate" at 566,2 size 50x50; CaptionText 'SIMATIC'
      on Change: "CheckDiagState"()
      ProcessValue <- "@DiagnosticsIndicatorTag"
   TextField "txtTitleBar" at 16,8 size 495x32; Text 'Application Name / Applikation'
   GraphicView "gfxNavigationIcon" at 1241,15 size 23x19; Picture "Hamburger_Icon"
   Button "btnNavigation" at 1224,0 size 56x48; TextOff 'Text'
      on Click: function_cf6f4242("GraphX_Slidein_Right", 1)
   IOField "Template_I/O field_1" at 1079,72 size 96x32; FormatPattern 9999999999999999999999999999999999999999
      ProcessValue <- "FB_LocalTime_DB_DateAndTIME"
   TextField "txtStateHeadline" at 75,55 size 123x23; Text 'State / Status'
   TextField "txtRecipeHeadline" at 281,55 size 154x23; Text 'Current Recipe / Rezeptur'
   TextField "txtOperatorHeadline" at 527,55 size 129x23; Text 'Operator / Bediener'
   SymbolicIOField "ioState" at 75,72 size 119x30; TextOn '1'; TextOff '0'; TextList "Machine State"
      ProcessValue <- "CurrentMachineState"
   IOField "ioRecipe" at 281,72 size 158x30; FormatPattern ??????????????????????????????
      ProcessValue <- "CurrentRecipeName"
   IOField "ioOperator" at 527,72 size 126x30; FormatPattern ??????????????????
      ProcessValue <- "CurrentUserName"
   Button "btnState" at 202,56 size 40x40; TextOff '...'; PictureOff "More_Icon"
      on Click: "ShowOperatingModePopUp"()
   Button "btnRecipe" at 449,56 size 40x40; TextOff '...'; PictureOff "More_Icon"
      on Click: "ShowRecipePopUp"()
   Rectangle "rectState" at 0,48 size 56x56
      Appearance <- "CurrentMachineState"
   Rectangle "rectSystemDiagnosticsIndicator" at 1224,48 size 56x56
      Appearance <- "DiagState"
   GraphicIOField "gioDiagState" at 1236,60 size 32x32; PictureList "DiagState_3"
      ProcessValue <- "DiagState"
   Button "btnDiagState" at 1224,48 size 56x56; TextOff 'Text'
      on Click: ActivateScreen("30_Diagnostics", 0)
   Button "btnOperator" at 669,56 size 40x40; TextOff '...'; PictureOff "More_Icon"
      on Click: "ShowLoginPopUp"()
   TextField "txtOperatorHeadline_1" at 768,55 size 129x23; Text 'Date and Time / Bediener'
   Button "btnOperator_1" at 995,56 size 40x40; TextOff '...'; PictureOff "More_Icon"
   DateTimeField "Template_Date/time field_1" at 768,72 size 208x30
      ProcessValue <- "FB_LocalTime_DB_DateAndTIME"
   Button "btnStartscreen" at 0,0 size 250x45; TextOff 'Text'
      on Click: "ActivateStartScreen"()
   Button "btnSubNavActive1" at 0,752 size 144x48; TextOff 'Overview / Übersicht'
      Visibility <- "SubNavigationState"
   Button "btnSubNavActive2" at 144,752 size 144x48; TextOff 'Module 1 / Modul 1'
      Visibility <- "SubNavigationState"
   Button "btnSubNavActive3" at 288,752 size 144x48; TextOff 'Module 2 / Modul 2'
      Visibility <- "SubNavigationState"
   Button "btnSubNavActive4" at 432,752 size 144x48; TextOff 'Module 3 / Modul 3'
      Visibility <- "SubNavigationState"
   Button "btnSubNavActive5" at 576,752 size 144x48; TextOff 'Module 4 / Modul 4'
      Visibility <- "SubNavigationState"
   Button "btnSubNavActive6" at 720,752 size 144x48; TextOff 'Module 5 / Modul 5'
      Visibility <- "SubNavigationState"
   Button "btnSubNavActive7" at 864,752 size 144x48; TextOff 'Module 6 / Modul 5'
      Visibility <- "SubNavigationState"
   Rectangle "rectIndicatorActive1" at 0,795 size 144x5
      Visibility <- "SubNavigationState"
   Rectangle "rectIndicatorActive2" at 144,795 size 144x5
      Visibility <- "SubNavigationState"
   Rectangle "rectIndicatorActive3" at 288,795 size 144x5
      Visibility <- "SubNavigationState"
   Rectangle "rectIndicatorActive4" at 432,795 size 144x5
      Visibility <- "SubNavigationState"
   Rectangle "rectIndicatorActive5" at 576,795 size 144x5
      Visibility <- "SubNavigationState"
   Rectangle "rectIndicatorActive6" at 720,795 size 144x5
      Visibility <- "SubNavigationState"
   Rectangle "rectIndicatorActive7" at 864,795 size 144x5
      Visibility <- "SubNavigationState"

Template "02_Two_Nav_Levels_Large_Text" 1280x800
   TextField "txtNextBackup1" at 16,120 size 232x24; Text 'Option 1'
   IOField "ioTargetPath1" at 16,152 size 236x24; FormatPattern ??????????????????????????????????????????????????
   TextField "txtNextBackup2" at 16,228 size 232x24; Text 'Option 2 / Option 1'
   IOField "ioTargetPath2" at 16,260 size 236x24; FormatPattern ??????????????????????????????????????????????????
   TextField "txtNextBackup3" at 16,336 size 232x24; Text 'Option 3 / Option 1'
   IOField "ioTargetPath3" at 16,368 size 236x24; FormatPattern ??????????????????????????????????????????????????
   TextField "txtNextBackup4" at 16,443 size 232x24; Text 'Option 4 / Option 1'
   IOField "ioTargetPath4" at 16,475 size 236x24; FormatPattern ??????????????????????????????????????????????????
   TextField "txtNextBackup5" at 16,551 size 232x24; Text 'Option 5 / Option 1'
   IOField "ioTargetPath5" at 16,583 size 236x24; FormatPattern ??????????????????????????????????????????????????
   TextField "txtNextBackup6" at 16,659 size 232x24; Text 'Option 6 / Option 1'
   IOField "ioTargetPath6" at 16,691 size 236x24; FormatPattern ??????????????????????????????????????????????????
   Button "btnSubNavigation1" at 0,104 size 264x109; TextOff 'Text'
      on Click: SetTag("ThirdLevelNavigationState", 1)
   Button "btnSubNavigation2" at 0,212 size 264x109; TextOff 'Text'
      on Click: SetTag("ThirdLevelNavigationState", 2)
   Button "btnSubNavigation3" at 0,320 size 264x109; TextOff 'Text'
      on Click: SetTag("ThirdLevelNavigationState", 3)
   Button "btnSubNavigation4" at 0,428 size 264x109; TextOff 'Text'
      on Click: SetTag("ThirdLevelNavigationState", 4)
   Button "btnSubNavigation5" at 0,536 size 264x109; TextOff 'Text'
      on Click: SetTag("ThirdLevelNavigationState", 5)
   Button "btnSubNavigation6" at 0,644 size 264x109; TextOff 'Text'
      on Click: SetTag("ThirdLevelNavigationState", 6)
   Gauge "gaugeDiagStateUpdate" at 566,2 size 50x50; CaptionText 'SIMATIC'
      on Change: "CheckDiagState"()
      ProcessValue <- "@DiagnosticsIndicatorTag"
   TextField "txtTitleBar" at 16,8 size 495x32; Text 'Packaging Machine / Applikation'
   GraphicView "gfxNavigationIcon" at 1241,15 size 23x19; Picture "Hamburger_Icon"
   Button "btnNavigation" at 1224,0 size 56x48; TextOff 'Text'
      on Click: function_cf6f4242("GraphX_Slidein_Right", 1)
   Button "btnStartscreen" at 0,0 size 250x45; TextOff 'Text'
      on Click: "ActivateStartScreen"()
   TextField "txtStateHeadline" at 75,55 size 123x23; Text 'State / Status'
   TextField "txtRecipeHeadline" at 281,55 size 154x23; Text 'Current Recipe / Rezeptur'
   TextField "txtOperatorHeadline" at 527,55 size 129x23; Text 'Operator / Bediener'
   SymbolicIOField "ioState" at 75,72 size 119x30; TextOn '1'; TextOff '0'; TextList "Machine State"
      ProcessValue <- "CurrentMachineState"
   IOField "ioRecipe" at 281,72 size 158x30; FormatPattern ??????????????????????????????
      ProcessValue <- "CurrentRecipeName"
   IOField "ioOperator" at 527,72 size 126x30; FormatPattern ??????????????????
      ProcessValue <- "CurrentUserName"
   Button "btnState" at 202,56 size 40x40; TextOff '...'; PictureOff "More_Icon"
      on Click: "ShowOperatingModePopUp"()
   Button "btnRecipe" at 449,56 size 40x40; TextOff '...'; PictureOff "More_Icon"
      on Click: "ShowRecipePopUp"()
   Rectangle "rectState" at 0,48 size 56x56
      Appearance <- "CurrentMachineState"
   Rectangle "rectSystemDiagnosticsIndicator" at 1224,48 size 56x56
      Appearance <- "DiagState"
   GraphicIOField "gioDiagState" at 1236,60 size 32x32; PictureList "DiagState_3"
      ProcessValue <- "DiagState"
   Button "btnDiagState" at 1224,48 size 56x56; TextOff 'Text'
      on Click: ActivateScreen("30_Diagnostics", 0)
   Button "btnOperator" at 669,56 size 40x40; TextOff '...'; PictureOff "More_Icon"
      on Click: "ShowLoginPopUp"()
   TextField "txtOperatorHeadline_1" at 768,55 size 129x23; Text 'Date and Time / Bediener'
   Button "btnOperator_1" at 995,56 size 40x40; TextOff '...'; PictureOff "More_Icon"
   DateTimeField "Template_Date/time field_1" at 768,72 size 208x30
   Rectangle "rectSubNavigation1" at 0,104 size 264x109
      Appearance <- "ThirdLevelNavigationState"
   Rectangle "rectSubNavigation2" at 0,212 size 264x109
      Appearance <- "ThirdLevelNavigationState"
   Rectangle "rectSubNavigation3" at 0,320 size 264x109
      Appearance <- "ThirdLevelNavigationState"
   Rectangle "rectSubNavigation4" at 0,428 size 264x109
      Appearance <- "ThirdLevelNavigationState"
   GraphicView "gfxPrevScreenIcon" at 1240,763 size 24x24; Picture "PrevScreen_Icon"
   Button "btnPreviousScreen" at 1224,751 size 56x48; TextOff 'Text'
      on Click: function_efd93a16()
   TextField "txtCurrentStateInfo" at 16,764 size 505x24; Text 'Optional Text about current state / Optionaler text mit aktuellem Status'
   Rectangle "rectSubNavigation4_1" at 0,536 size 264x109
      Appearance <- "ThirdLevelNavigationState"
   Rectangle "rectSubNavigation4_2" at 0,644 size 264x108
      Appearance <- "ThirdLevelNavigationState"

Template "02_Two_Nav_Levels_Text" 1280x800
   Button "btnSubNav1" at 0,146 size 144x56; TextOn 'Item 1'; TextOff 'Item 1'
      on Click: SetTag("SubNavigationState", 1)
   Button "btnSubNav2" at 0,201 size 144x56; TextOn 'Item 2'; TextOff 'Item 2'
      on Click: SetTag("SubNavigationState", 2)
   Button "btnSubNav3" at 0,256 size 144x60; TextOn 'Item 3'; TextOff 'Item 3'
      on Click: SetTag("SubNavigationState", 3)
   Button "btnSubNav4" at 0,315 size 144x60; TextOn 'Item 4'; TextOff 'Item 4'
      on Click: SetTag("SubNavigationState", 4)
   Button "btnSubNav5" at 0,374 size 144x60; TextOn 'Item 5'; TextOff 'Item 5'
      on Click: SetTag("SubNavigationState", 4)
   GraphicView "gfxRuntimeStop" at 61,763 size 23x28; Picture "Power_dark"
   Button "btnRuntimeStop" at 0,752 size 144x48; TextOff 'Text'
      on Click: StopRuntime(0)
   Button "btnSubNavActive1" at 0,146 size 144x56; TextOff 'Item 1 / Display'
      Visibility <- "SubNavigationState"
   Button "btnSubNavActive2" at 0,201 size 144x56; TextOff 'Item 2'
      Visibility <- "SubNavigationState"
   Button "btnSubNavActive3" at 0,256 size 144x60; TextOff 'Item 3'
      Visibility <- "SubNavigationState"
   Button "btnSubNavActive4" at 0,315 size 144x60; TextOff 'Item 4'
      Visibility <- "SubNavigationState"
   Button "btnSubNavActive5" at 0,374 size 144x60; TextOn 'Item 5'; TextOff 'Item 5'
      Visibility <- "SubNavigationState"
   Rectangle "rectIndicatorActive1" at 0,146 size 5x56
      Visibility <- "SubNavigationState"
   Rectangle "rectIndicatorActive2" at 0,201 size 5x56
      Visibility <- "SubNavigationState"
   Rectangle "rectIndicatorActive3" at 0,256 size 5x60
      Visibility <- "SubNavigationState"
   Rectangle "rectIndicatorActive4" at 0,315 size 5x60
      Visibility <- "SubNavigationState"
   Rectangle "rectIndicatorActive5" at 0,374 size 5x60
      Visibility <- "SubNavigationState"
   Gauge "gaugeDiagStateUpdate" at 566,2 size 50x50; CaptionText 'SIMATIC'
      on Change: "CheckDiagState"()
      ProcessValue <- "@DiagnosticsIndicatorTag"
   TextField "txtTitleBar" at 16,8 size 495x32; Text 'Application Name / Applikation'
   GraphicView "gfxNavigationIcon" at 1241,15 size 23x19; Picture "Hamburger_Icon"
   Button "btnNavigation" at 1224,0 size 56x48; TextOff 'Text'
      on Click: function_cf6f4242("GraphX_Slidein_Right", 1)
   Button "btnStartscreen" at 0,0 size 250x45; TextOff 'Text'
      on Click: "ActivateStartScreen"()
   TextField "txtStateHeadline" at 75,55 size 123x23; Text 'State / Status'
   TextField "txtRecipeHeadline" at 281,55 size 154x23; Text 'Current Recipe / Rezeptur'
   TextField "txtOperatorHeadline" at 527,55 size 129x23; Text 'Operator / Bediener'
   SymbolicIOField "ioState" at 75,72 size 119x30; TextOn '1'; TextOff '0'; TextList "Machine State"
      ProcessValue <- "CurrentMachineState"
   IOField "ioRecipe" at 281,72 size 158x30; FormatPattern ??????????????????????????????
      ProcessValue <- "CurrentRecipeName"
   IOField "ioOperator" at 527,72 size 126x30; FormatPattern ??????????????????
      ProcessValue <- "CurrentUserName"
   Button "btnState" at 202,56 size 40x40; TextOff '...'; PictureOff "More_Icon"
      on Click: "ShowOperatingModePopUp"()
   Button "btnRecipe" at 449,56 size 40x40; TextOff '...'; PictureOff "More_Icon"
      on Click: "ShowRecipePopUp"()
   Rectangle "rectState" at 0,48 size 56x56
      Appearance <- "CurrentMachineState"
   Rectangle "rectSystemDiagnosticsIndicator" at 1224,48 size 56x56
      Appearance <- "DiagState"
   GraphicIOField "gioDiagState" at 1236,60 size 32x32; PictureList "DiagState_3"
      ProcessValue <- "DiagState"
   Button "btnDiagState" at 1224,48 size 56x56; TextOff 'Text'
      on Click: ActivateScreen("30_Diagnostics", 0)
   Button "btnOperator" at 669,56 size 40x40; TextOff '...'; PictureOff "More_Icon"
      on Click: "ShowLoginPopUp"()
   TextField "txtOperatorHeadline_1" at 768,55 size 129x23; Text 'Date and Time / Bediener'
   Button "btnOperator_1" at 995,56 size 40x40; TextOff '...'; PictureOff "More_Icon"
   DateTimeField "Template_Date/time field_1" at 768,72 size 208x30